(* Logix 5000 project; controller Almacen_1 vendor 1 type 14 code 235 rev 36.11; software revision 36.00 *) (continued)
   T_Permissive_HomeStep2 : TIMER;
   T_Permissive_HomeStep3 : TIMER;
   T_Permissive_HomeStep4 : TIMER;
   T_Permissive_HomeStep5 : TIMER;
   T_Permissive_HomeStep6 : TIMER;
   T_Permissive_HomeStep7 : TIMER;
   T_Permissive_HomeStep8 : TIMER;
   T_Permissive_HomeStep9 : TIMER;
   T_Permissive_HomStep0 : TIMER;
   T_Pieza_Antes_Marcadora : TIMER;
   T_Pieza_Camara : TIMER;
   T_Pieza_FinDeCarrera : TIMER;
   T_Pieza_FinDeCarrera_Error : TIMER;
   T_Pieza_FinDeCarrera_Salida : TIMER;
   T_Pieza_Marcadora : TIMER;
   T_Pieza_MarcadoraTerminada : TIMER;
   T_Pieza_TomaFanuc : TIMER;
   Test_Bit : DINT := 537136129;
   Timer_1 : TIMER;
   Timer_2 : TIMER;
   Timer_3 : TIMER;
   Timer_4 : TIMER;
   Timer_5 : TIMER;
   Timer_6 : TIMER;
   Timer_7 : TIMER;
   Timer_8 : TIMER;
   To_Pos_Alm_1 : DINT := 64; {produced}
   Tope_CNC_Conv_1 : BOOL;   // Tope Pistón CNC (Freno 5) Conveyor 1
   Tope_CNC_Conv_2 : BOOL;   // Tope Pistón CNC (Freno 5) Conveyor 2
   Tope_Marcadora_Conv_1 : BOOL;   // Tope Pistón Marcadora Láser (Freno 6) Conveyor 1
   Tope_Marcadora_Conv_2 : BOOL;   // Tope Pistón Marcadora Láser (Freno 6) Conveyor 2
   Tope_Salida_PH_Conv_1 : BOOL;   // Tope Pistón Salida de Producto (Freno 8) Conveyor 1
   Tope_Salida_PH_Conv_2 : BOOL;   // Tope Pistón Salida de Producto (Freno 8) Conveyor 2
   Tope_Vision_Conv_1 : BOOL;   // Tope Pistón Cáma de Visión Conveyor 1
   Tope_Vision_Conv_2 : BOOL;   // Tope Pistón Cámara de Visión Conveyor 2
   Usar_Proceso_CNC_1_de_Conveyor_1 : BOOL;   // Bit Para usar pasos del Robot Fanuc en el Conveyor 1
   X_Negative : BOOL;
   X_Positive : BOOL := 1;
   Y_Negative : BOOL := 1;
   Y_Positive : BOOL;
   Yaw_Negative : BOOL := 1;
   Yaw_Positive : BOOL;
   Yellow_Light_Alm_1 : BOOL := 1;
   Yellow_Light_Alm_2 : BOOL;
END_VAR

PROGRAM _02_Conveyor_1
VAR
   CamOnline : BOOL := 1;
   CompletedNS : BOOL;
   Count1 : COUNTER;
   Inspecting : BOOL;
   JobPass : BOOL;
   Timer : TIMER; {access Read Only}
   Timer1 : TIMER;
   Timer2 : TIMER;
   Timer3 : TIMER;
   Timer5 : TIMER; {access Read Only}
   trigger : BOOL := 1;
   TriggerGus1 : BOOL;
   TriggerGusEN : BOOL := 1;
   Valid : BOOL;
END_VAR
END_PROGRAM

PROGRAM MainProgram   (* main routine MainRoutine *)
VAR
   Contador : COUNTER;
   Contador_Salida_Conveyor : COUNTER;
   End_Conveyor_Rutine : BOOL;
   mem1 : BOOL;
   mem2 : BOOL;
   mem3 : BOOL;
   mem4 : BOOL;
   mem5 : BOOL;
   PosDer_Alm_0_C : BOOL;
   PosDer_Alm_0_E : BOOL;
   PosDer_Alm_1_C : BOOL;
   PosDer_Alm_1_E : BOOL;
   PosDer_Alm_2_C : BOOL;
   PosDer_Alm_2_E : BOOL;
   PosDer_Alm_3_C : BOOL;
   PosDer_Alm_3_E : BOOL;
   PosDer_Alm_4_C : BOOL;
   PosDer_Alm_4_E : BOOL;
   PosDer_Alm_5_C : BOOL;
   PosDer_Alm_5_E : BOOL;
   PosIzq_Alm_0_C : BOOL;
   PosIzq_Alm_0_E : BOOL;
   PosIzq_Alm_1_C : BOOL;
   PosIzq_Alm_1_E : BOOL;
   PosIzq_Alm_2_C : BOOL;
   PosIzq_Alm_2_E : BOOL;
   PosIzq_Alm_3_C : BOOL;
   PosIzq_Alm_3_E : BOOL;
   PosIzq_Alm_4_C : BOOL;
   PosIzq_Alm_4_E : BOOL;
   PosIzq_Alm_5_C : BOOL;
   PosIzq_Alm_5_E : BOOL;
   PosIzq_Alm_6_C : BOOL;
   PosIzq_Conv_6_C : BOOL;
   PosIzq_Conv_8_C : BOOL;
   PosIzq_Conv_8_E : BOOL;
   PosProgramming : BOOL;
   Start_Conveyor_1 : BOOL;
   Start_Rutine : BOOL := 1;
   Stop_Conveyor_1 : BOOL;
   tag_switch : BOOL;
   tag_switch2 : BOOL;
   tag_switch3 : BOOL;
   Tag_switch4 : BOOL;
   tag_switch5 : BOOL;
   tag_switch6 : BOOL;
   tag_timer_piston : BOOL;
   tag_timer_piston2 : BOOL;
   TEMP1 : TIMER;
   TIM2 : TIMER;
   TIM3 : TIMER;
   TIM4 : TIMER;
   Timer1_Cambio_Direccion_CNC : TIMER;
   Timer2 : TIMER;
   Timer3_Piston_Marcadora_OFF : TIMER;
   Timer4_Piston_Camara_ON : TIMER;
   Timer5_Piston_Camara_OFF : TIMER;
   Timer6_Cambio_Direccion_Almacen : TIMER;
   Timer7_Sensor_Entrada_Salida : TIMER;
   Timer8_Stop_Conveyor : TIMER;
   Timer9_Piston_Salida : TIMER;
END_VAR

ROUTINE Almacen1   (* ladder *)
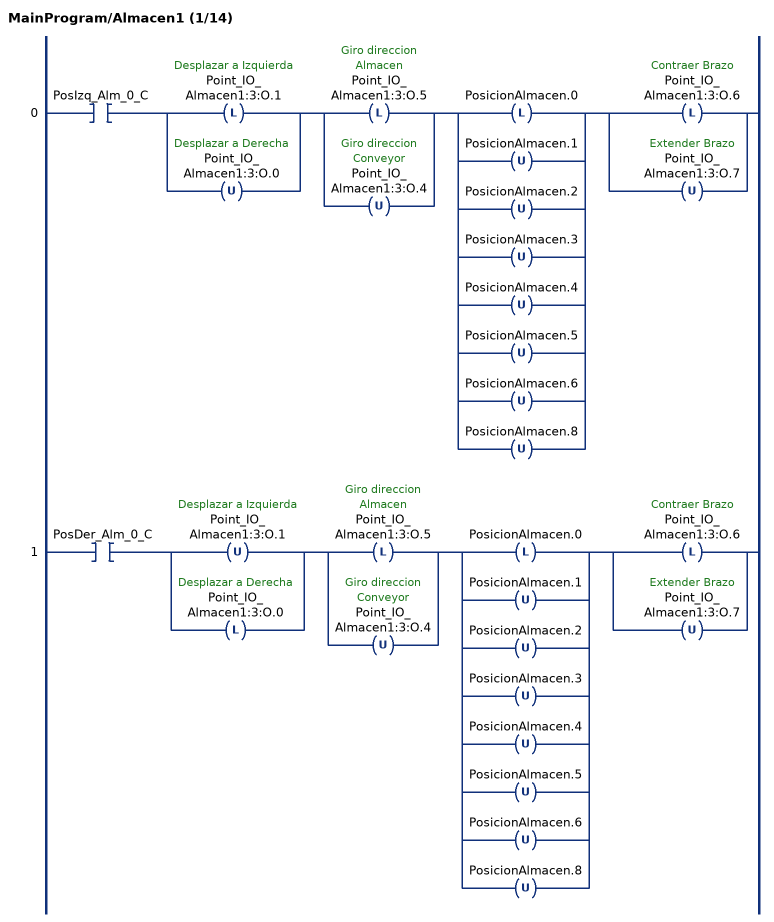
   0: XIC(PosIzq_Alm_0_C)[OTL(Point_IO_Almacen1:3:O.1) ,OTU(Point_IO_Almacen1:3:O.0) ][OTL(Point_IO_Almacen1:3:O.5) ,OTU(Point_IO_Almacen1:3:O.4) ][OTL(PosicionAlmacen.0) ,OTU(PosicionAlmacen.1) ,OTU(PosicionAlmacen.2) ,OTU(PosicionAlmacen.3) ,OTU(PosicionAlmacen.4) ,OTU(PosicionAlmacen.5) ,OTU(PosicionAlmacen.6) ,OTU(PosicionAlmacen.8) ][OTL(Point_IO_Almacen1:3:O.6) ,OTU(Point_IO_Almacen1:3:O.7) ];
   1: XIC(PosDer_Alm_0_C)[OTU(Point_IO_Almacen1:3:O.1) ,OTL(Point_IO_Almacen1:3:O.0) ][OTL(Point_IO_Almacen1:3:O.5) ,OTU(Point_IO_Almacen1:3:O.4) ][OTL(PosicionAlmacen.0) ,OTU(PosicionAlmacen.1) ,OTU(PosicionAlmacen.2) ,OTU(PosicionAlmacen.3) ,OTU(PosicionAlmacen.4) ,OTU(PosicionAlmacen.5) ,OTU(PosicionAlmacen.6) ,OTU(PosicionAlmacen.8) ][OTL(Point_IO_Almacen1:3:O.6) ,OTU(Point_IO_Almacen1:3:O.7) ];
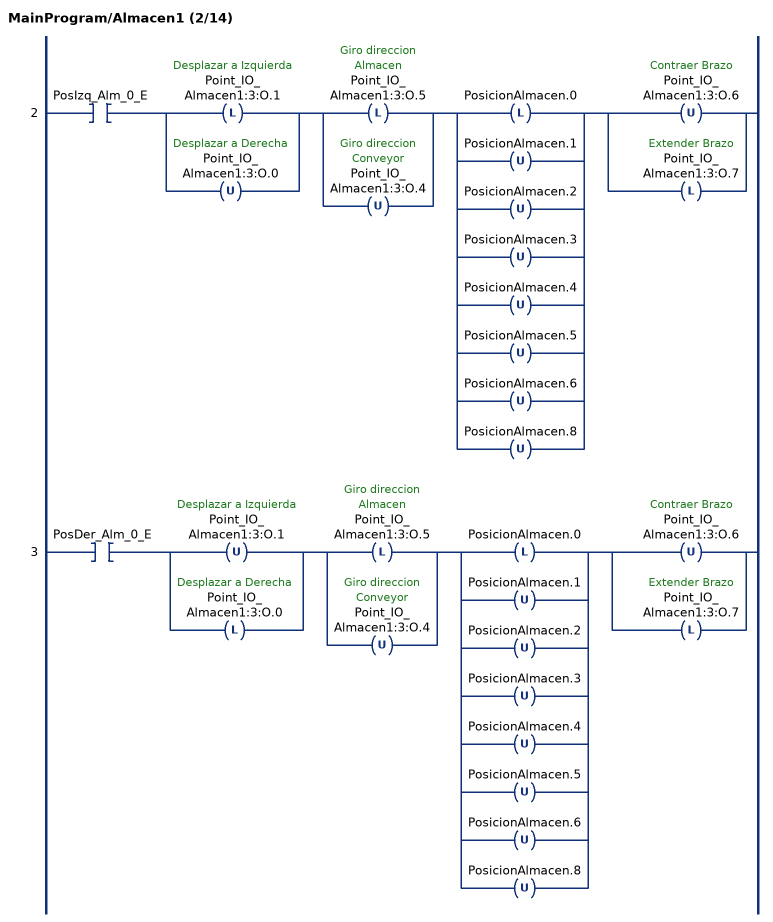
   2: XIC(PosIzq_Alm_0_E)[OTL(Point_IO_Almacen1:3:O.1) ,OTU(Point_IO_Almacen1:3:O.0) ][OTL(Point_IO_Almacen1:3:O.5) ,OTU(Point_IO_Almacen1:3:O.4) ][OTL(PosicionAlmacen.0) ,OTU(PosicionAlmacen.1) ,OTU(PosicionAlmacen.2) ,OTU(PosicionAlmacen.3) ,OTU(PosicionAlmacen.4) ,OTU(PosicionAlmacen.5) ,OTU(PosicionAlmacen.6) ,OTU(PosicionAlmacen.8) ][OTU(Point_IO_Almacen1:3:O.6) ,OTL(Point_IO_Almacen1:3:O.7) ];
   3: XIC(PosDer_Alm_0_E)[OTU(Point_IO_Almacen1:3:O.1) ,OTL(Point_IO_Almacen1:3:O.0) ][OTL(Point_IO_Almacen1:3:O.5) ,OTU(Point_IO_Almacen1:3:O.4) ][OTL(PosicionAlmacen.0) ,OTU(PosicionAlmacen.1) ,OTU(PosicionAlmacen.2) ,OTU(PosicionAlmacen.3) ,OTU(PosicionAlmacen.4) ,OTU(PosicionAlmacen.5) ,OTU(PosicionAlmacen.6) ,OTU(PosicionAlmacen.8) ][OTU(Point_IO_Almacen1:3:O.6) ,OTL(Point_IO_Almacen1:3:O.7) ];
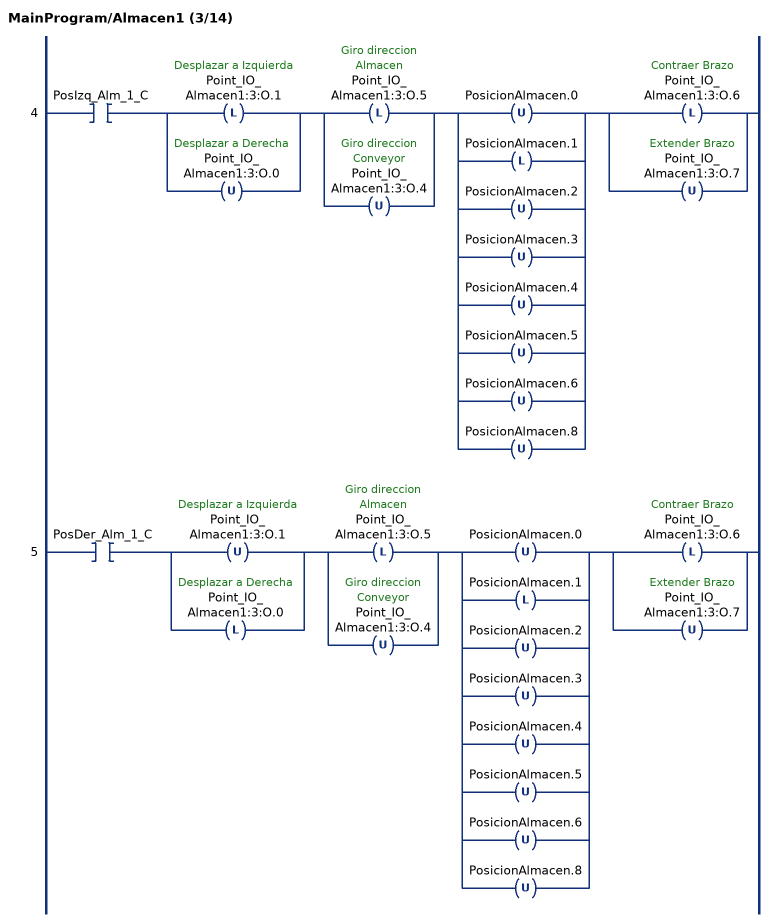
   4: XIC(PosIzq_Alm_1_C)[OTL(Point_IO_Almacen1:3:O.1) ,OTU(Point_IO_Almacen1:3:O.0) ][OTL(Point_IO_Almacen1:3:O.5) ,OTU(Point_IO_Almacen1:3:O.4) ][OTU(PosicionAlmacen.0) ,OTL(PosicionAlmacen.1) ,OTU(PosicionAlmacen.2) ,OTU(PosicionAlmacen.3) ,OTU(PosicionAlmacen.4) ,OTU(PosicionAlmacen.5) ,OTU(PosicionAlmacen.6) ,OTU(PosicionAlmacen.8) ][OTL(Point_IO_Almacen1:3:O.6) ,OTU(Point_IO_Almacen1:3:O.7) ];
   5: XIC(PosDer_Alm_1_C)[OTU(Point_IO_Almacen1:3:O.1) ,OTL(Point_IO_Almacen1:3:O.0) ][OTL(Point_IO_Almacen1:3:O.5) ,OTU(Point_IO_Almacen1:3:O.4) ][OTU(PosicionAlmacen.0) ,OTL(PosicionAlmacen.1) ,OTU(PosicionAlmacen.2) ,OTU(PosicionAlmacen.3) ,OTU(PosicionAlmacen.4) ,OTU(PosicionAlmacen.5) ,OTU(PosicionAlmacen.6) ,OTU(PosicionAlmacen.8) ][OTL(Point_IO_Almacen1:3:O.6) ,OTU(Point_IO_Almacen1:3:O.7) ];
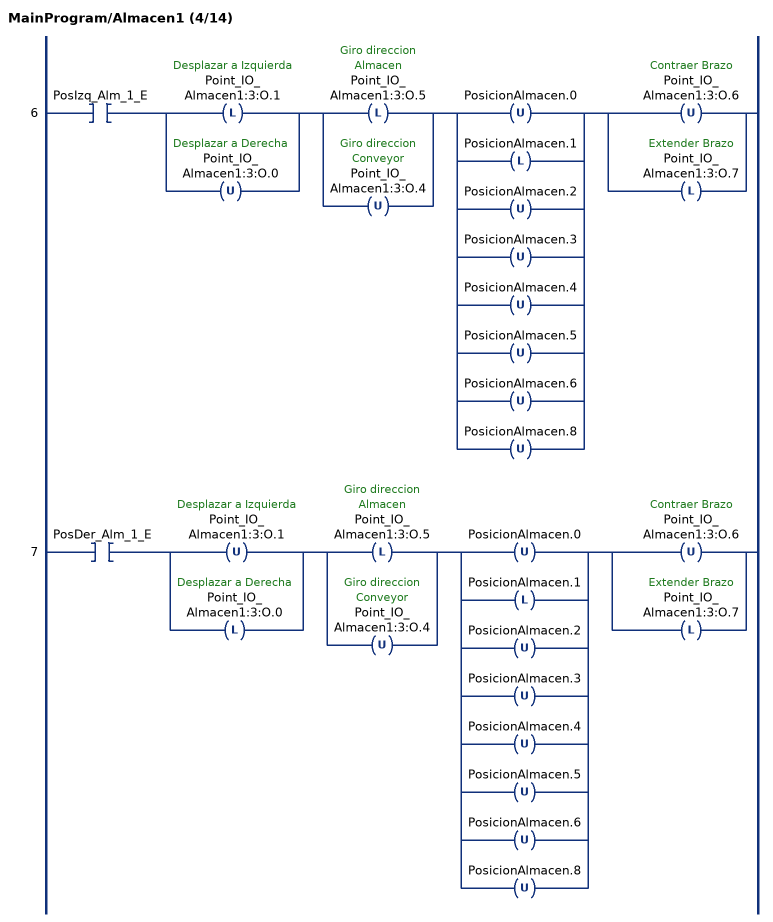
   6: XIC(PosIzq_Alm_1_E)[OTL(Point_IO_Almacen1:3:O.1) ,OTU(Point_IO_Almacen1:3:O.0) ][OTL(Point_IO_Almacen1:3:O.5) ,OTU(Point_IO_Almacen1:3:O.4) ][OTU(PosicionAlmacen.0) ,OTL(PosicionAlmacen.1) ,OTU(PosicionAlmacen.2) ,OTU(PosicionAlmacen.3) ,OTU(PosicionAlmacen.4) ,OTU(PosicionAlmacen.5) ,OTU(PosicionAlmacen.6) ,OTU(PosicionAlmacen.8) ][OTU(Point_IO_Almacen1:3:O.6) ,OTL(Point_IO_Almacen1:3:O.7) ];
   7: XIC(PosDer_Alm_1_E)[OTU(Point_IO_Almacen1:3:O.1) ,OTL(Point_IO_Almacen1:3:O.0) ][OTL(Point_IO_Almacen1:3:O.5) ,OTU(Point_IO_Almacen1:3:O.4) ][OTU(PosicionAlmacen.0) ,OTL(PosicionAlmacen.1) ,OTU(PosicionAlmacen.2) ,OTU(PosicionAlmacen.3) ,OTU(PosicionAlmacen.4) ,OTU(PosicionAlmacen.5) ,OTU(PosicionAlmacen.6) ,OTU(PosicionAlmacen.8) ][OTU(Point_IO_Almacen1:3:O.6) ,OTL(Point_IO_Almacen1:3:O.7) ];
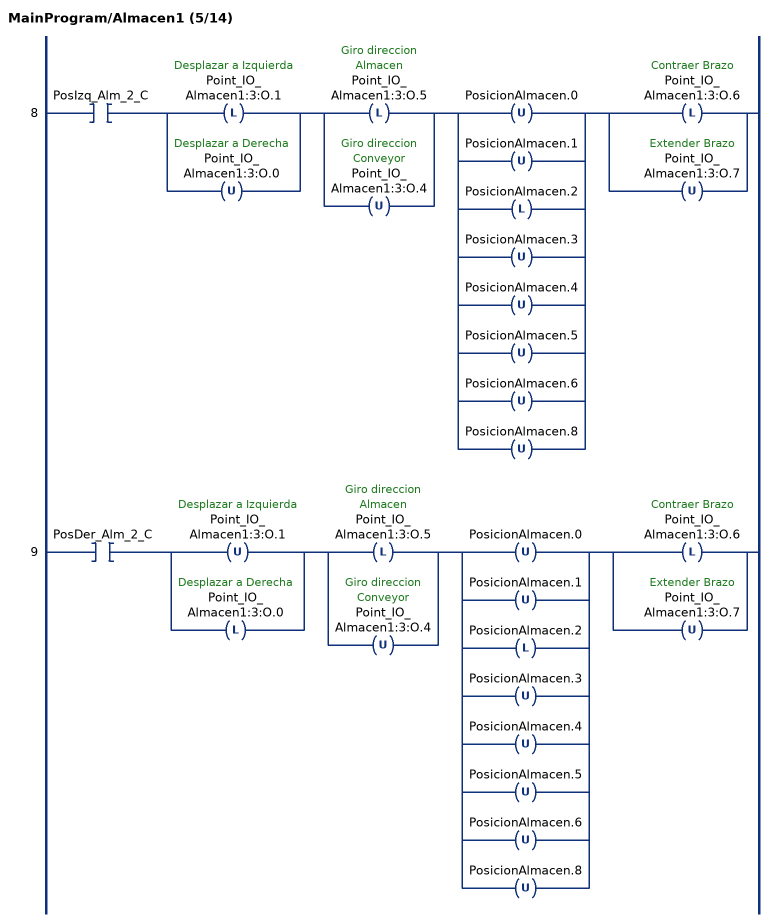
   8: XIC(PosIzq_Alm_2_C)[OTL(Point_IO_Almacen1:3:O.1) ,OTU(Point_IO_Almacen1:3:O.0) ][OTL(Point_IO_Almacen1:3:O.5) ,OTU(Point_IO_Almacen1:3:O.4) ][OTU(PosicionAlmacen.0) ,OTU(PosicionAlmacen.1) ,OTL(PosicionAlmacen.2) ,OTU(PosicionAlmacen.3) ,OTU(PosicionAlmacen.4) ,OTU(PosicionAlmacen.5) ,OTU(PosicionAlmacen.6) ,OTU(PosicionAlmacen.8) ][OTL(Point_IO_Almacen1:3:O.6) ,OTU(Point_IO_Almacen1:3:O.7) ];
   9: XIC(PosDer_Alm_2_C)[OTU(Point_IO_Almacen1:3:O.1) ,OTL(Point_IO_Almacen1:3:O.0) ][OTL(Point_IO_Almacen1:3:O.5) ,OTU(Point_IO_Almacen1:3:O.4) ][OTU(PosicionAlmacen.0) ,OTU(PosicionAlmacen.1) ,OTL(PosicionAlmacen.2) ,OTU(PosicionAlmacen.3) ,OTU(PosicionAlmacen.4) ,OTU(PosicionAlmacen.5) ,OTU(PosicionAlmacen.6) ,OTU(PosicionAlmacen.8) ][OTL(Point_IO_Almacen1:3:O.6) ,OTU(Point_IO_Almacen1:3:O.7) ];
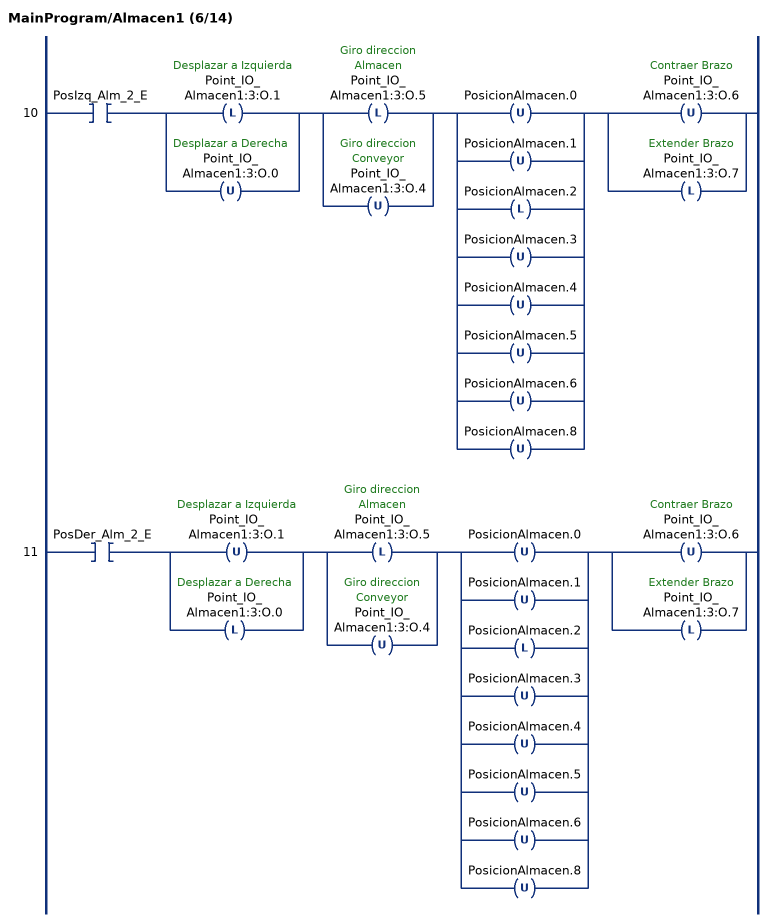
   10: XIC(PosIzq_Alm_2_E)[OTL(Point_IO_Almacen1:3:O.1) ,OTU(Point_IO_Almacen1:3:O.0) ][OTL(Point_IO_Almacen1:3:O.5) ,OTU(Point_IO_Almacen1:3:O.4) ][OTU(PosicionAlmacen.0) ,OTU(PosicionAlmacen.1) ,OTL(PosicionAlmacen.2) ,OTU(PosicionAlmacen.3) ,OTU(PosicionAlmacen.4) ,OTU(PosicionAlmacen.5) ,OTU(PosicionAlmacen.6) ,OTU(PosicionAlmacen.8) ][OTU(Point_IO_Almacen1:3:O.6) ,OTL(Point_IO_Almacen1:3:O.7) ];
   11: XIC(PosDer_Alm_2_E)[OTU(Point_IO_Almacen1:3:O.1) ,OTL(Point_IO_Almacen1:3:O.0) ][OTL(Point_IO_Almacen1:3:O.5) ,OTU(Point_IO_Almacen1:3:O.4) ][OTU(PosicionAlmacen.0) ,OTU(PosicionAlmacen.1) ,OTL(PosicionAlmacen.2) ,OTU(PosicionAlmacen.3) ,OTU(PosicionAlmacen.4) ,OTU(PosicionAlmacen.5) ,OTU(PosicionAlmacen.6) ,OTU(PosicionAlmacen.8) ][OTU(Point_IO_Almacen1:3:O.6) ,OTL(Point_IO_Almacen1:3:O.7) ];
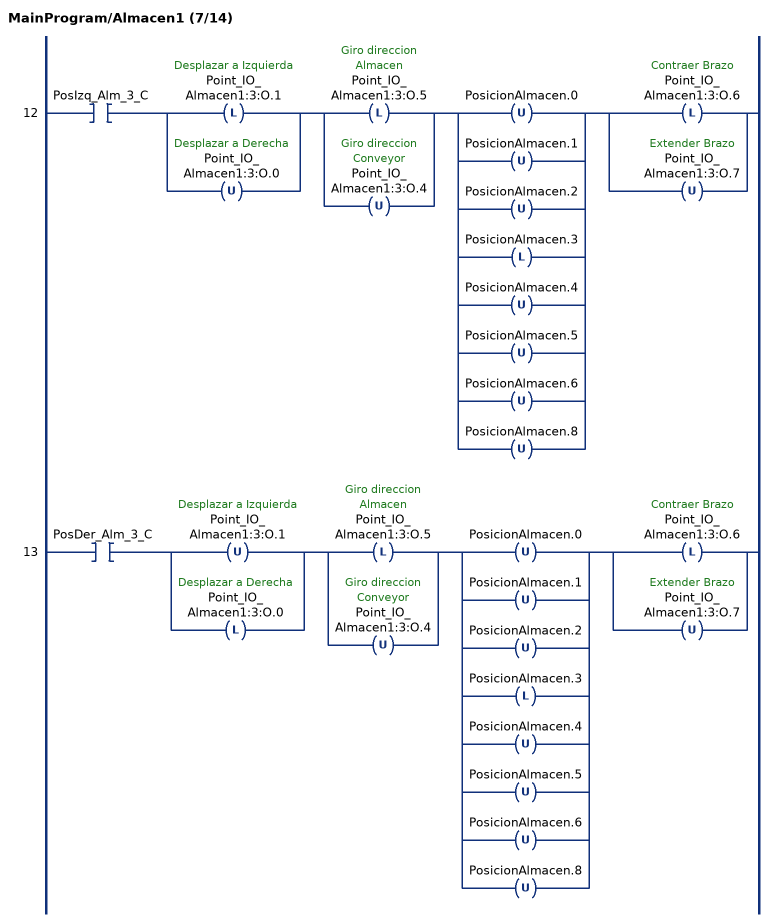
   12: XIC(PosIzq_Alm_3_C)[OTL(Point_IO_Almacen1:3:O.1) ,OTU(Point_IO_Almacen1:3:O.0) ][OTL(Point_IO_Almacen1:3:O.5) ,OTU(Point_IO_Almacen1:3:O.4) ][OTU(PosicionAlmacen.0) ,OTU(PosicionAlmacen.1) ,OTU(PosicionAlmacen.2) ,OTL(PosicionAlmacen.3) ,OTU(PosicionAlmacen.4) ,OTU(PosicionAlmacen.5) ,OTU(PosicionAlmacen.6) ,OTU(PosicionAlmacen.8) ][OTL(Point_IO_Almacen1:3:O.6) ,OTU(Point_IO_Almacen1:3:O.7) ];
   13: XIC(PosDer_Alm_3_C)[OTU(Point_IO_Almacen1:3:O.1) ,OTL(Point_IO_Almacen1:3:O.0) ][OTL(Point_IO_Almacen1:3:O.5) ,OTU(Point_IO_Almacen1:3:O.4) ][OTU(PosicionAlmacen.0) ,OTU(PosicionAlmacen.1) ,OTU(PosicionAlmacen.2) ,OTL(PosicionAlmacen.3) ,OTU(PosicionAlmacen.4) ,OTU(PosicionAlmacen.5) ,OTU(PosicionAlmacen.6) ,OTU(PosicionAlmacen.8) ][OTL(Point_IO_Almacen1:3:O.6) ,OTU(Point_IO_Almacen1:3:O.7) ];
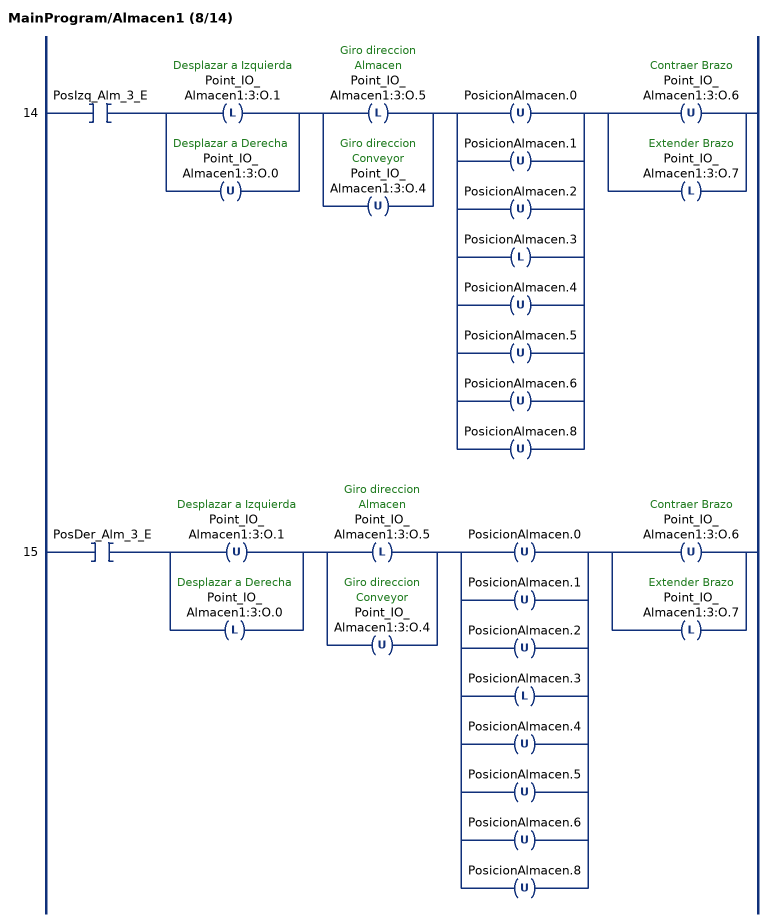
   14: XIC(PosIzq_Alm_3_E)[OTL(Point_IO_Almacen1:3:O.1) ,OTU(Point_IO_Almacen1:3:O.0) ][OTL(Point_IO_Almacen1:3:O.5) ,OTU(Point_IO_Almacen1:3:O.4) ][OTU(PosicionAlmacen.0) ,OTU(PosicionAlmacen.1) ,OTU(PosicionAlmacen.2) ,OTL(PosicionAlmacen.3) ,OTU(PosicionAlmacen.4) ,OTU(PosicionAlmacen.5) ,OTU(PosicionAlmacen.6) ,OTU(PosicionAlmacen.8) ][OTU(Point_IO_Almacen1:3:O.6) ,OTL(Point_IO_Almacen1:3:O.7) ];
   15: XIC(PosDer_Alm_3_E)[OTU(Point_IO_Almacen1:3:O.1) ,OTL(Point_IO_Almacen1:3:O.0) ][OTL(Point_IO_Almacen1:3:O.5) ,OTU(Point_IO_Almacen1:3:O.4) ][OTU(PosicionAlmacen.0) ,OTU(PosicionAlmacen.1) ,OTU(PosicionAlmacen.2) ,OTL(PosicionAlmacen.3) ,OTU(PosicionAlmacen.4) ,OTU(PosicionAlmacen.5) ,OTU(PosicionAlmacen.6) ,OTU(PosicionAlmacen.8) ][OTU(Point_IO_Almacen1:3:O.6) ,OTL(Point_IO_Almacen1:3:O.7) ];
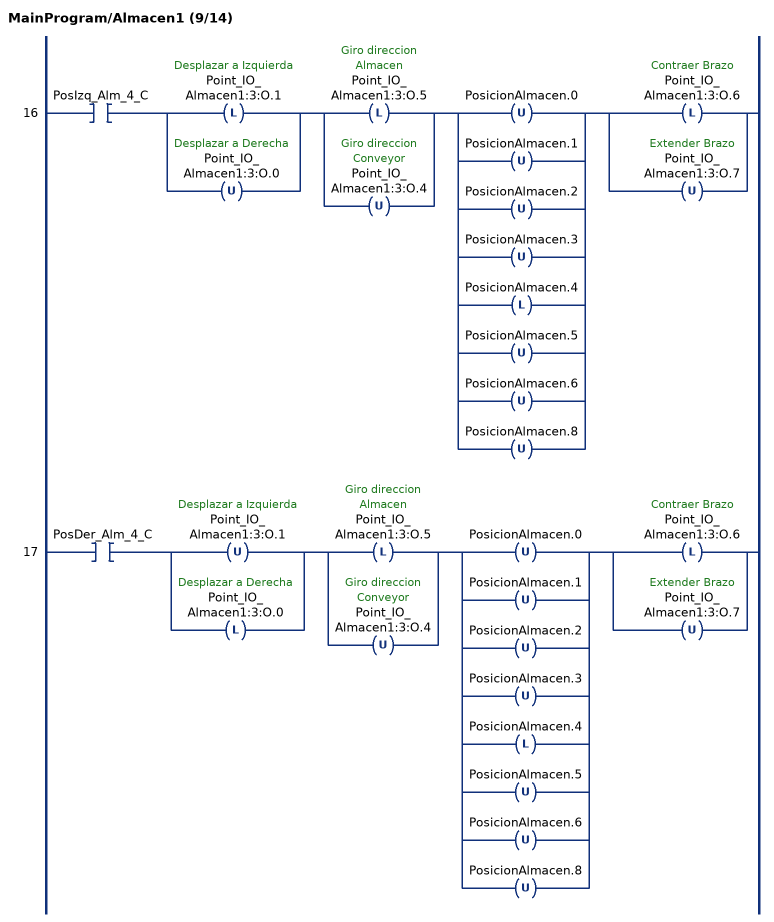
   16: XIC(PosIzq_Alm_4_C)[OTL(Point_IO_Almacen1:3:O.1) ,OTU(Point_IO_Almacen1:3:O.0) ][OTL(Point_IO_Almacen1:3:O.5) ,OTU(Point_IO_Almacen1:3:O.4) ][OTU(PosicionAlmacen.0) ,OTU(PosicionAlmacen.1) ,OTU(PosicionAlmacen.2) ,OTU(PosicionAlmacen.3) ,OTL(PosicionAlmacen.4) ,OTU(PosicionAlmacen.5) ,OTU(PosicionAlmacen.6) ,OTU(PosicionAlmacen.8) ][OTL(Point_IO_Almacen1:3:O.6) ,OTU(Point_IO_Almacen1:3:O.7) ];
   17: XIC(PosDer_Alm_4_C)[OTU(Point_IO_Almacen1:3:O.1) ,OTL(Point_IO_Almacen1:3:O.0) ][OTL(Point_IO_Almacen1:3:O.5) ,OTU(Point_IO_Almacen1:3:O.4) ][OTU(PosicionAlmacen.0) ,OTU(PosicionAlmacen.1) ,OTU(PosicionAlmacen.2) ,OTU(PosicionAlmacen.3) ,OTL(PosicionAlmacen.4) ,OTU(PosicionAlmacen.5) ,OTU(PosicionAlmacen.6) ,OTU(PosicionAlmacen.8) ][OTL(Point_IO_Almacen1:3:O.6) ,OTU(Point_IO_Almacen1:3:O.7) ];
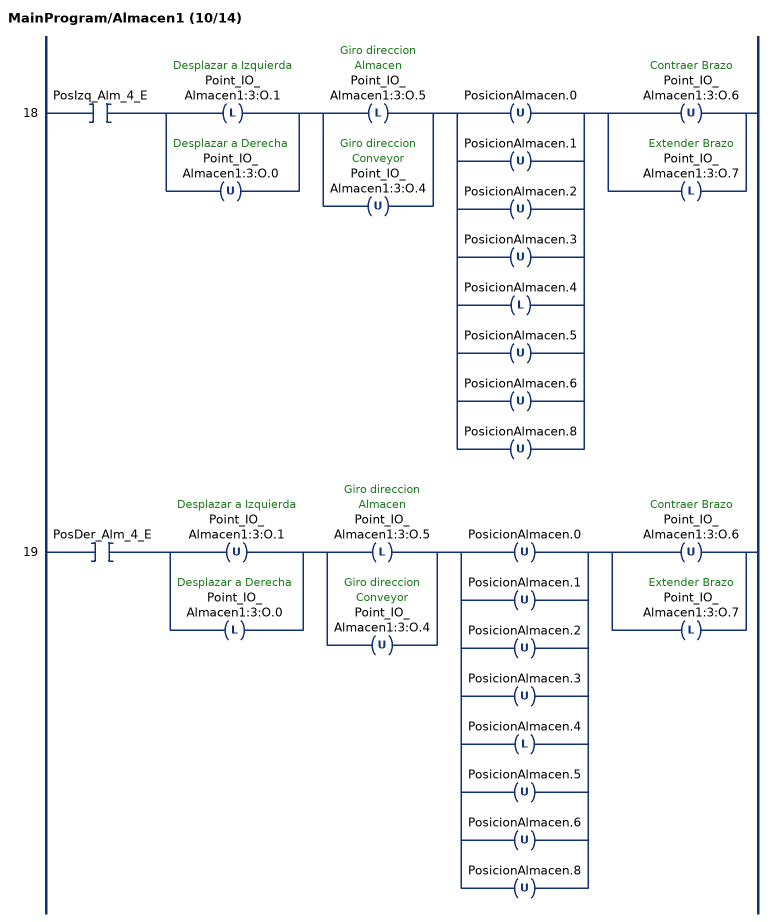
   18: XIC(PosIzq_Alm_4_E)[OTL(Point_IO_Almacen1:3:O.1) ,OTU(Point_IO_Almacen1:3:O.0) ][OTL(Point_IO_Almacen1:3:O.5) ,OTU(Point_IO_Almacen1:3:O.4) ][OTU(PosicionAlmacen.0) ,OTU(PosicionAlmacen.1) ,OTU(PosicionAlmacen.2) ,OTU(PosicionAlmacen.3) ,OTL(PosicionAlmacen.4) ,OTU(PosicionAlmacen.5) ,OTU(PosicionAlmacen.6) ,OTU(PosicionAlmacen.8) ][OTU(Point_IO_Almacen1:3:O.6) ,OTL(Point_IO_Almacen1:3:O.7) ];
   19: XIC(PosDer_Alm_4_E)[OTU(Point_IO_Almacen1:3:O.1) ,OTL(Point_IO_Almacen1:3:O.0) ][OTL(Point_IO_Almacen1:3:O.5) ,OTU(Point_IO_Almacen1:3:O.4) ][OTU(PosicionAlmacen.0) ,OTU(PosicionAlmacen.1) ,OTU(PosicionAlmacen.2) ,OTU(PosicionAlmacen.3) ,OTL(PosicionAlmacen.4) ,OTU(PosicionAlmacen.5) ,OTU(PosicionAlmacen.6) ,OTU(PosicionAlmacen.8) ][OTU(Point_IO_Almacen1:3:O.6) ,OTL(Point_IO_Almacen1:3:O.7) ];
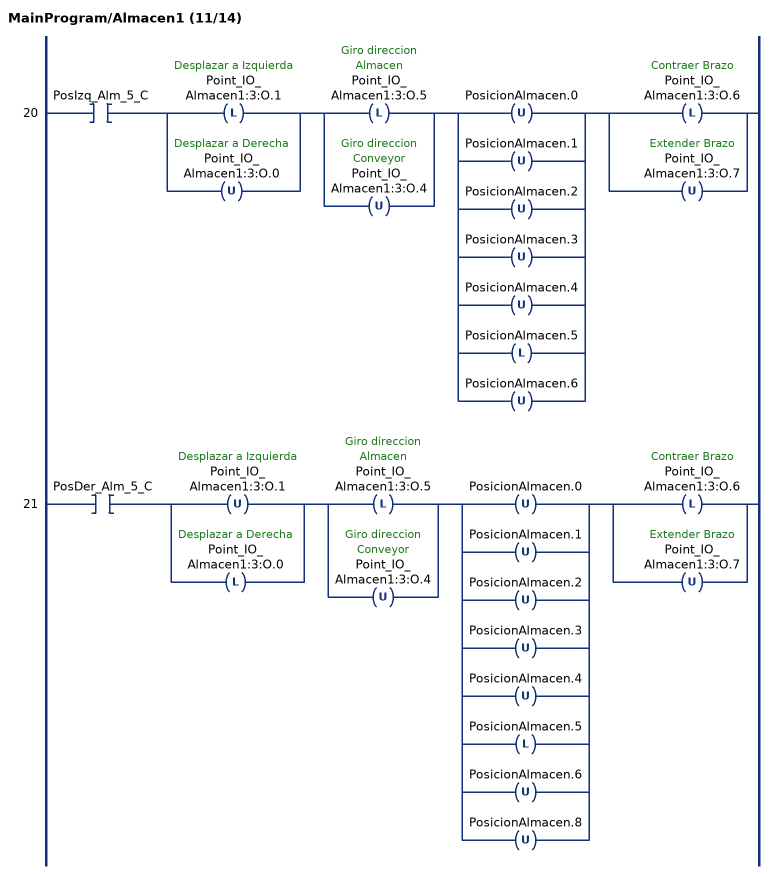
   20: XIC(PosIzq_Alm_5_C)[OTL(Point_IO_Almacen1:3:O.1) ,OTU(Point_IO_Almacen1:3:O.0) ][OTL(Point_IO_Almacen1:3:O.5) ,OTU(Point_IO_Almacen1:3:O.4) ][OTU(PosicionAlmacen.0) ,OTU(PosicionAlmacen.1) ,OTU(PosicionAlmacen.2) ,OTU(PosicionAlmacen.3) ,OTU(PosicionAlmacen.4) ,OTL(PosicionAlmacen.5) ,OTU(PosicionAlmacen.6) ][OTL(Point_IO_Almacen1:3:O.6) ,OTU(Point_IO_Almacen1:3:O.7) ];
   21: XIC(PosDer_Alm_5_C)[OTU(Point_IO_Almacen1:3:O.1) ,OTL(Point_IO_Almacen1:3:O.0) ][OTL(Point_IO_Almacen1:3:O.5) ,OTU(Point_IO_Almacen1:3:O.4) ][OTU(PosicionAlmacen.0) ,OTU(PosicionAlmacen.1) ,OTU(PosicionAlmacen.2) ,OTU(PosicionAlmacen.3) ,OTU(PosicionAlmacen.4) ,OTL(PosicionAlmacen.5) ,OTU(PosicionAlmacen.6) ,OTU(PosicionAlmacen.8) ][OTL(Point_IO_Almacen1:3:O.6) ,OTU(Point_IO_Almacen1:3:O.7) ];
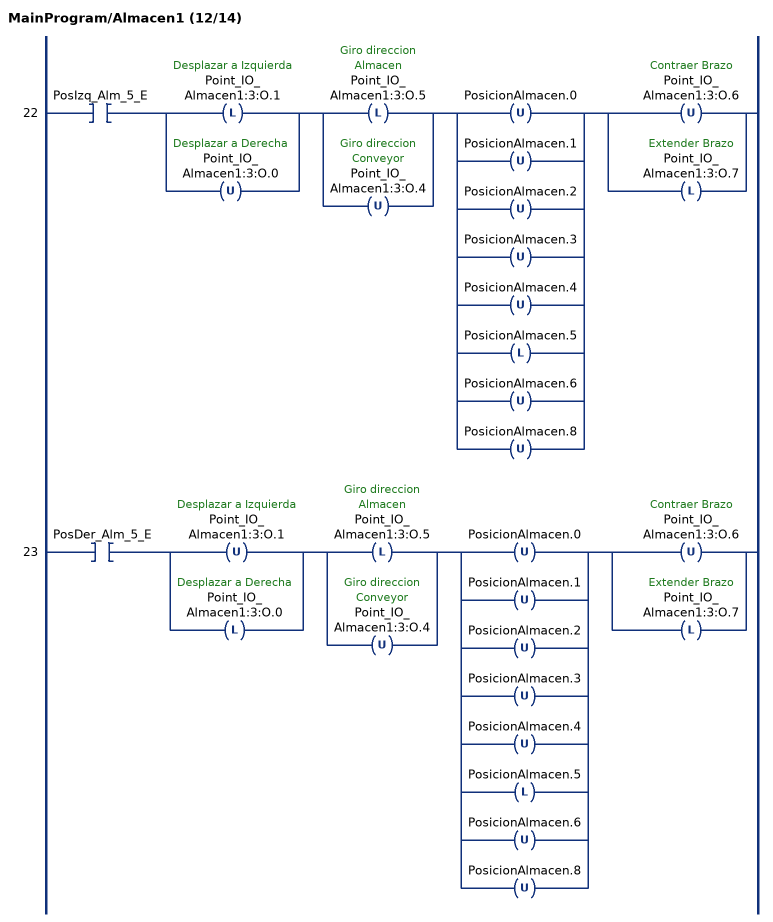
   22: XIC(PosIzq_Alm_5_E)[OTL(Point_IO_Almacen1:3:O.1) ,OTU(Point_IO_Almacen1:3:O.0) ][OTL(Point_IO_Almacen1:3:O.5) ,OTU(Point_IO_Almacen1:3:O.4) ][OTU(PosicionAlmacen.0) ,OTU(PosicionAlmacen.1) ,OTU(PosicionAlmacen.2) ,OTU(PosicionAlmacen.3) ,OTU(PosicionAlmacen.4) ,OTL(PosicionAlmacen.5) ,OTU(PosicionAlmacen.6) ,OTU(PosicionAlmacen.8) ][OTU(Point_IO_Almacen1:3:O.6) ,OTL(Point_IO_Almacen1:3:O.7) ];
   23: XIC(PosDer_Alm_5_E)[OTU(Point_IO_Almacen1:3:O.1) ,OTL(Point_IO_Almacen1:3:O.0) ][OTL(Point_IO_Almacen1:3:O.5) ,OTU(Point_IO_Almacen1:3:O.4) ][OTU(PosicionAlmacen.0) ,OTU(PosicionAlmacen.1) ,OTU(PosicionAlmacen.2) ,OTU(PosicionAlmacen.3) ,OTU(PosicionAlmacen.4) ,OTL(PosicionAlmacen.5) ,OTU(PosicionAlmacen.6) ,OTU(PosicionAlmacen.8) ][OTU(Point_IO_Almacen1:3:O.6) ,OTL(Point_IO_Almacen1:3:O.7) ];
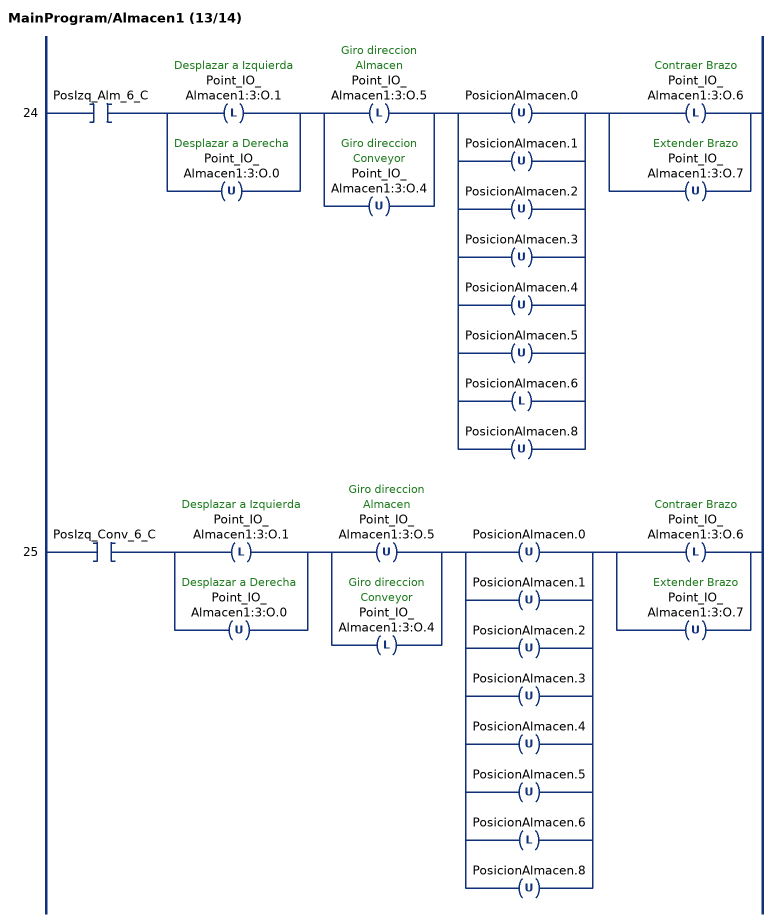
   24: XIC(PosIzq_Alm_6_C)[OTL(Point_IO_Almacen1:3:O.1) ,OTU(Point_IO_Almacen1:3:O.0) ][OTL(Point_IO_Almacen1:3:O.5) ,OTU(Point_IO_Almacen1:3:O.4) ][OTU(PosicionAlmacen.0) ,OTU(PosicionAlmacen.1) ,OTU(PosicionAlmacen.2) ,OTU(PosicionAlmacen.3) ,OTU(PosicionAlmacen.4) ,OTU(PosicionAlmacen.5) ,OTL(PosicionAlmacen.6) ,OTU(PosicionAlmacen.8) ][OTL(Point_IO_Almacen1:3:O.6) ,OTU(Point_IO_Almacen1:3:O.7) ];
   25: XIC(PosIzq_Conv_6_C)[OTL(Point_IO_Almacen1:3:O.1) ,OTU(Point_IO_Almacen1:3:O.0) ][OTU(Point_IO_Almacen1:3:O.5) ,OTL(Point_IO_Almacen1:3:O.4) ][OTU(PosicionAlmacen.0) ,OTU(PosicionAlmacen.1) ,OTU(PosicionAlmacen.2) ,OTU(PosicionAlmacen.3) ,OTU(PosicionAlmacen.4) ,OTU(PosicionAlmacen.5) ,OTL(PosicionAlmacen.6) ,OTU(PosicionAlmacen.8) ][OTL(Point_IO_Almacen1:3:O.6) ,OTU(Point_IO_Almacen1:3:O.7) ];
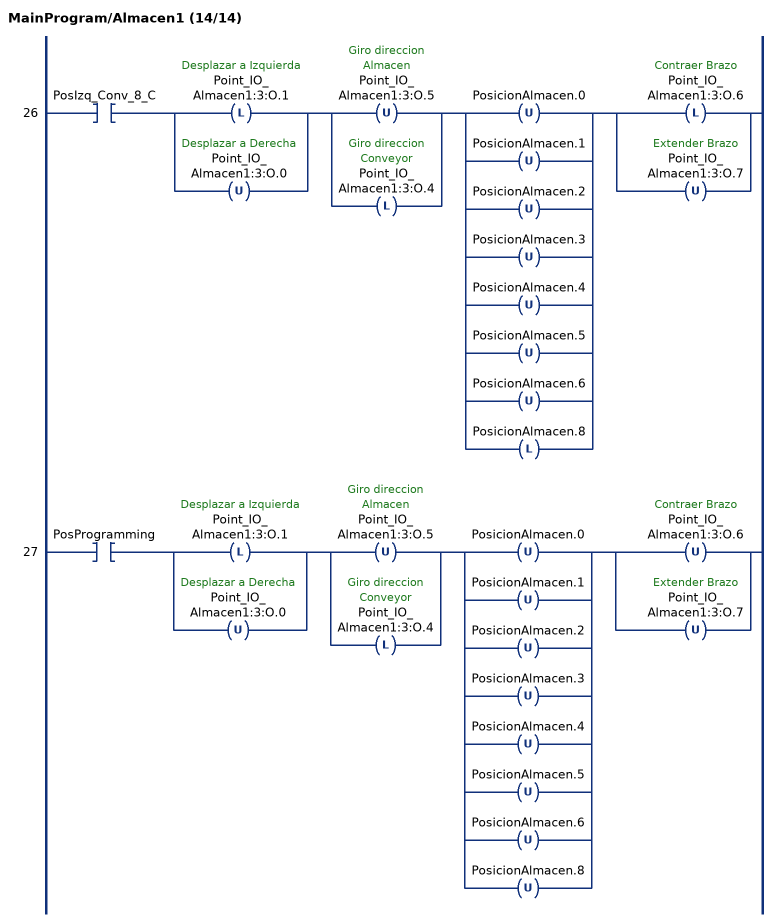
   26: XIC(PosIzq_Conv_8_C)[OTL(Point_IO_Almacen1:3:O.1) ,OTU(Point_IO_Almacen1:3:O.0) ][OTU(Point_IO_Almacen1:3:O.5) ,OTL(Point_IO_Almacen1:3:O.4) ][OTU(PosicionAlmacen.0) ,OTU(PosicionAlmacen.1) ,OTU(PosicionAlmacen.2) ,OTU(PosicionAlmacen.3) ,OTU(PosicionAlmacen.4) ,OTU(PosicionAlmacen.5) ,OTU(PosicionAlmacen.6) ,OTL(PosicionAlmacen.8) ][OTL(Point_IO_Almacen1:3:O.6) ,OTU(Point_IO_Almacen1:3:O.7) ];
   27: XIC(PosProgramming)[OTL(Point_IO_Almacen1:3:O.1) ,OTU(Point_IO_Almacen1:3:O.0) ][OTU(Point_IO_Almacen1:3:O.5) ,OTL(Point_IO_Almacen1:3:O.4) ][OTU(PosicionAlmacen.0) ,OTU(PosicionAlmacen.1) ,OTU(PosicionAlmacen.2) ,OTU(PosicionAlmacen.3) ,OTU(PosicionAlmacen.4) ,OTU(PosicionAlmacen.5) ,OTU(PosicionAlmacen.6) ,OTU(PosicionAlmacen.8) ][OTU(Point_IO_Almacen1:3:O.6) ,OTU(Point_IO_Almacen1:3:O.7) ];
END_ROUTINE
